           IF (#iSP <> #old.SP // SP has changed.
               OR #RTIRG_auto.Q // Auto has just been enabled, and the valve is out of pos.
               (* *)AND ABS(#iSP - #io.in.pos) > #conf.regModeMinOffset
               OR NOT #iMan AND ( // In auto
               (* *)#RTIRG_iReset.Q // Avoid dead lock
               (* *)OR #RTRIG_iFailSafe_released.Q
               (* *)OR #RTRIG_iInterlook_released.Q
               (* *)OR #RTRIG_jogClose_released.Q OR #RTRIG_jogOpen_released.Q )
               (* *)) AND (
               (*     *)NOT #iRegMode // Not regMode, no aditional requirements.
               (*     *)OR #TON_regModeWait.Q AND ( // A break between each move.
               (*        *)// Offset is bigger then a certain offset.
               (*        *)ABS(#iSP - #io.in.pos) > #conf.regModeMinOffset
               (*        *)// At almost closed and open, the offset requirement
               (*        *)// may not be fulfilled.
               (*        *)OR #io.in.pos > #conf.fullyOpenPosLim - #conf.endPosWithoutPreStop
               (*        *)OR #io.in.pos < #conf.endPosWithoutPreStop))
               // regMode should be used when a valve is controlled by a PID.
               // When the valve is in regMode, then there will be a time break between each 
               // movment. And there is a need a certain offset before an ajustment is done.
               // This behavior significantly prevents wear on the valve. If the valve is not
               // in regMode, then each change in SP will make the valve operate.
           THEN
               IF #iSP > #io.in.pos THEN
                   #action := #OPEN;
               ELSIF #iSP < #io.in.pos THEN
                   #action := #CLOSE;
               END_IF;
           END_IF;

           // --------------------------------------
           // SP-reached-pos:
           // 
           // In the main area where the valve operate, it will shut off the outputs, a
           // tiny bit before it reach the SP. This make the valve, stop exacly on SP.
           // In the area of almost closed and almost open this function is disable,
           // this makes sure that it's possible to open or close the valve entirly.
           #pre := SEL(G := #iSP > #conf.fullyOpenPosLim - #conf.endPosWithoutPreStop
                       OR #iSP < #conf.endPosWithoutPreStop,
                       IN0 := #conf.preStop, IN1 := 0);
           // Detect reached position
           IF #action = #OPEN AND (#io.in.pos > #iSP - #pre OR #io.in.fullyOpen)
               OR #action = #CLOSE AND (#io.in.pos < #iSP + #pre OR #io.in.fullyClosed)
           THEN
               #action := #NO_ACTION;
               RESET_TIMER(#TON_regModeWait);
           END_IF;
       END_IF;
       // In regMode this timer need to finnish before a new movement can be done.
       #TON_regModeWait.TON(IN := true,
                            PT := #conf.regModeTimeBreak);
   END_REGION

   REGION Gentle
       // If a big valve closes or open to fast, it can damage the pipes or other
       // equipment. This section make time breaks on closing or opening. 

       #gentleMode := #io.in.pos < #conf.gentleActivteLowLimit // ->
       // -> The function is only active under a ceratain position limit.
       AND (NOT #iFailSafe OR #conf.gentleAlsoOnFailSafe)
       // AlsoOnFailSafe: It's possible to disable the function for emergencies
       // by setting the value false.
       AND (#conf.gentleOpenEnable AND #action = #OPEN
       (* *)OR #conf.gentleCloseEnable AND #action = #CLOSE);    

       // The time break will increase as the valve move from the limit towards close.
       #pause := REAL_TO_DINT(#conf.gentleTimePauseBias
                              + (#io.in.pos / #conf.gentleActivteLowLimit)
                              * #conf.gentleTimePauseDelta);
       IF #gentleMode THEN
           #TON_gentle.TON(IN := true,
                           PT := SEL(G := #gentleAction, // Toggle times
                                     IN0 := #conf.gentleTimeRun,
                                     IN1 := #pause));
           IF #TON_gentle.Q THEN
               #gentleAction := NOT #gentleAction;
               RESET_TIMER(#TON_gentle); 
           END_IF;
           #action2 := SEL(G := #gentleAction, // Toggle action
                           IN0 := #action, IN1 := #NO_ACTION);
       ELSE
           RESET_TIMER(#TON_gentle);
           #gentleAction := false;
           // If the carefully-function is disabled, then just forward
           // the action value to the next stage.
           #action2 := #action;
       END_IF;
   END_REGION

   REGION Output
       // Make a smal time break when valve change direction. This make sure that
       // that both outputs are not active at the same time.
       #TP_toggleOut.TP(IN := #action2 <> #old.action2 AND #old.action2 <> #NO_ACTION,
                        PT := #conf.toggleTimeBreak);

       // Outputs
       IF #TP_toggleOut.Q THEN // A small time break.
           #io.out.open := false;
           #io.out.close := false;
       ELSIF #iFailSafe 
           OR #iJogClose OR #iJogOpen
       THEN
           // When failSafe or jog is active both the limit-switch and positon
           // signal most indicate that the valve is in correct position. This
           // in case one of the signals isn't working.
           #io.out.open := #action2 = #OPEN AND NOT #bothSensors.open;
           #io.out.close := #action2 = #CLOSE AND NOT #bothSensors.closed;
       ELSIF #iInterlook THEN
           #io.out.open := false;
           #io.out.close := false;
       ELSE
           #io.out.open := #action2 = #OPEN AND NOT #io.in.fullyOpen;
           #io.out.close := #action2 = #CLOSE AND NOT #io.in.fullyClosed;
       END_IF;
   END_REGION

   REGION Old    
       // Store values, to check if they has changed until next scan.
       #old.SP := #iSP;
       #old.action := #action;
       #old.action2 := #action2;
   END_REGION

   #qTimeout := #out.qucikTimeout OR #out.longTimeout;
END_FUNCTION_BLOCK

FUNCTION_BLOCK "motorValve"   // FB10, SCL
{ S7_Optimized_Access := 'TRUE' }
VERSION : 0.1
   VAR_INPUT
      iFeedbackPosition : Real;
      iFeddbackPosError : Bool;
      iFeedbackFullyOpen : Bool;
      iFeedbackFullyClosed : Bool;
   END_VAR
   VAR_OUTPUT
      qOpen : Bool;
      qClose : Bool := FALSE;
   END_VAR
   VAR RETAIN
      hmi : "motorValveHmiUdt";
   END_VAR
   VAR
      valve : "motorValveCtrl";
      SP : Real;
      SP_auto : Real;
   END_VAR
   VAR CONSTANT
      AUTO : SInt := 0;
      MAN_LOCAL : SInt := 1;
      MAN_REMOTE : SInt := 2;
   END_VAR
BEGIN
   // Valve with analog feedback.

   REGION Simulation
       IF #hmi.sim.enable AND NOT #valve.iFailSafe THEN
           // Simulation of input signal, not possible if in fail safe mode.
           #hmi.io.in.pos := #hmi.sim.pos;
           #hmi.io.in.posError := false;
           #hmi.io.in.fullyOpen := #hmi.sim.pos > #hmi.conf.fullyOpenPosLim;
           #hmi.io.in.fullyClosed := #hmi.sim.pos < #hmi.conf.fullyClosedPosLim;
       ELSE
           // Input mapping
           #hmi.io.in.pos := #iFeedbackPosition;
           #hmi.io.in.posError := #iFeddbackPosError;
           #hmi.io.in.fullyOpen := #iFeedbackFullyOpen;
           #hmi.io.in.fullyClosed := #iFeedbackFullyClosed;
       END_IF;
   END_REGION

   REGION Man / auto    
       IF #hmi.cmd.stop THEN
           #hmi.autoMan := #MAN_LOCAL;
       ELSIF #hmi.cmd.jogOpen XOR #hmi.cmd.jogClose THEN
           #hmi.autoMan := #MAN_LOCAL;
           #SP := #iFeedbackPosition;
       ELSIF #hmi.cmd.openFully XOR #hmi.cmd.closeFully THEN
           #hmi.autoMan := #MAN_LOCAL;
           #SP := SEL(G := #hmi.cmd.openFully, IN0 := 0, IN1 := 100);
       ELSIF #hmi.autoMan = #MAN_LOCAL THEN
           #SP := #hmi.SP;
       ELSIF #hmi.autoMan = #AUTO THEN
           #SP := #SP_auto;
           // If auto is controlled by a pid then #hmi.conf.regMode need to be enabled.
       END_IF;
       #hmi.SP := #valve.iSP := #SP_auto := #SP;
       // Forward auto or man to the valve controller.
       CASE #hmi.autoMan OF
           #MAN_LOCAL, #MAN_REMOTE:
               #valve.iMan := true;
           #AUTO:
               #valve.iMan := false;
       END_CASE;
   END_REGION

   REGION Valve controller.        
       // Main valve controller block.
       #valve(// iFailSafe
              // iInterlook
              // iRegMode
              iStop := #hmi.cmd.stop,
              iJogOpen := #hmi.cmd.jogOpen,
              iJogClose := #hmi.cmd.jogClose,
              iReset := #hmi.cmd.reset,
              qTimeout => #hmi.error.timeout,
              conf := #hmi.conf,
              io := #hmi.io);
       #qOpen := #hmi.io.out.open; // Outputs
       #qClose := #hmi.io.out.close;
   END_REGION

   REGION Position error    
       #hmi.error.posError :=
       #iFeedbackFullyOpen AND #iFeedbackFullyClosed
       OR #iFeedbackFullyOpen
       (* *)AND #iFeedbackPosition < #hmi.conf.fullyOpenPosLim - #hmi.conf.regModeMinOffset
       (* *)AND NOT #hmi.conf.simFullyOpenWithPos
       OR #iFeedbackFullyClosed
       (* *)AND #iFeedbackPosition > #hmi.conf.fullyClosedPosLim + #hmi.conf.regModeMinOffset
       (* *)AND NOT #hmi.conf.simFullyClosedWithPos;
   END_REGION

   REGION End
       // Count secounds the valve has been operating, and number of starts.
       "operatingTime"(in := #qOpen OR #qClose,
                       opr := #hmi.operatingTime);

       // Reset signals.
       #hmi.cmd.jogOpen := false;
       #hmi.cmd.jogClose := false;
       #hmi.cmd.openFully := false;
       #hmi.cmd.closeFully := false;
       #hmi.cmd.reset := false;
       #hmi.cmd.man := false;
       #hmi.cmd.auto := false;
       CASE #hmi.autoMan OF // Reset stop signal, only if in man.
           #MAN_LOCAL, #MAN_REMOTE: // If in auto, then do nothing.
               #hmi.cmd.stop := false;
       END_CASE;

       // Other signals to HMI
       #hmi.info.failSafe := #valve.iFailSafe;
       #hmi.info.interlook := #valve.iInterlook;
       #hmi.info.regMode := #valve.iRegMode;

       #hmi.sim.simByPlc := #hmi.io.simulated;
       #hmi.io.simulated := false;
   END_REGION
END_FUNCTION_BLOCK

FUNCTION_BLOCK "motorValveSimulation"   // FB20, SCL
{ S7_Optimized_Access := 'TRUE' }
VERSION : 0.1
   VAR_INPUT
      speed : Real := 1.0;
   END_VAR
   VAR_IN_OUT
      io : "motorValveIoUdt";
   END_VAR
   VAR
      old : UDInt;
      sn : UDInt;
   END_VAR
   VAR_TEMP
      t : DTL;
      "e" : Int;
   END_VAR
BEGIN
   #"e" := RD_SYS_T(#t);
   #sn := #t.NANOSECOND / 100000 + #t.SECOND * 10;

   IF #sn = #old THEN
       IF #io.out.open THEN
           #io.in.pos += #speed * 0.1;
       ELSIF #io.out.close THEN
           #io.in.pos -= #speed;
       END_IF;
   END_IF;
   #old := #sn;

   #io.in.pos := LIMIT(MN := 0, IN := #io.in.pos, MX := 100);
   #io.in.fullyOpen := #io.in.pos > 99;
   #io.in.fullyClosed := #io.in.pos < 1;

   #io.simulated := true;
END_FUNCTION_BLOCK

// folder: _ state macine

FUNCTION_BLOCK "stateMachineTimer"   // FB1, SCL
{ S7_Optimized_Access := 'TRUE' }
VERSION : 0.1
   VAR_INPUT
      state : Int;   // state machine
   END_VAR
   VAR_OUTPUT
      q : Bool;   // out
      rt : Time;   // Remaining time
      et : Time;
   END_VAR
   VAR
      pt : Time;   // input time
      "timer" : IEC_TIMER;
      old_state : Int;
   END_VAR
BEGIN
   // https://github.com/rexhip/
   //
   // State machine timer.
   // 
   // The timer is reseted if:
   // - Pt hasen't got a new value (for each scan)
   // - New state

   #"timer".TON(IN := #pt <> T#0s
              (* *)AND #state = #old_state,
              PT := #pt,
              Q => #q);

   #et := #"timer".ET;
   #rt := #pt - #et;

   #pt := T#0s;
   #old_state := #state;
END_FUNCTION_BLOCK

FUNCTION_BLOCK "setResetTimer"   // FB3, SCL
{ S7_Optimized_Access := 'TRUE' }
VERSION : 0.1
   VAR_INPUT
      in : Bool;
      pt : Time;
      set : Bool;
      reset : Bool;
   END_VAR
   VAR_OUTPUT
      q : Bool;
   END_VAR
   VAR
      "timer" : IEC_TIMER;
      timer_q : Bool;
   END_VAR
BEGIN
   // Once the timer has elapsed, the output
   // will stay true until it's reset.

   #"timer".TON(IN := #in, PT := #pt, Q => #timer_q);

   IF #set THEN
       #q := true;
   ELSIF #reset THEN
       #q := false;
   ELSIF #timer_q THEN
       #q := true;
   END_IF;
END_FUNCTION_BLOCK

FUNCTION "sTimer" : Bool   // FC2, SCL
{ S7_Optimized_Access := 'TRUE' }
VERSION : 0.1
   VAR_INPUT
      pt : Time;
   END_VAR
   VAR_IN_OUT
      t : "stateMachineTimer";
   END_VAR
BEGIN
   // sTimer
   // Make a timer, a one liner, in a state macine

   #t.pt := #pt;
   #sTimer := #t.q;
END_FUNCTION

// folder: io

FUNCTION_BLOCK "ioGlobal_FB"   // FB1, SCL
{ S7_Optimized_Access := 'TRUE' }
VERSION : 0.1
   VAR
      hmi : "ioGlobalUdt";
      z_internal_timer : IEC_TIMER;
      z_internal : Struct
         fs : Bool := TRUE;
         timer_mem : Time;
      END_STRUCT;
      collectInfo : Struct
         activeSimCnt : UInt;
         activeAlarmsCnt : UInt;
         unacknowledgedAlarmsCnt : UInt;
         errorCnt : UInt;
      END_STRUCT;
      info2ioBlocks : Struct
         runtimeDiff : Time;
         ackAllAlarms : Bool;
         disableAllSim : Bool;
         firstScan : Bool := TRUE;
      END_STRUCT;
      z : Struct
         ioIdCnt : UInt;
      END_STRUCT;
      copyPaste : "analogInAndAlarmsUdt";
      normX : "normXAnalogUdt";
   END_VAR
BEGIN
   // ioGlobal: This block handels common function for io, eg:
   //  - Count active simulations
   //  - Disable all simulations
   //  - Count active alarms
   //  - Ack. all active alarms

   // Calculate time of each plc scan.
   #z_internal_timer.TON(IN := NOT #z_internal_timer.Q, PT := T#24d);
   IF #z_internal_timer.ET <> #z_internal.timer_mem THEN
       #info2ioBlocks.runtimeDiff := #z_internal_timer.ET - #z_internal.timer_mem;
   END_IF;
   #z_internal.timer_mem := #z_internal_timer.ET;

   // First scan
   #info2ioBlocks.firstScan := #z_internal.fs;
   #z_internal.fs := false;

   // Common information to all io-blocks.
   #info2ioBlocks.ackAllAlarms := #hmi.ackAllAlarms;
   #info2ioBlocks.disableAllSim := #hmi.disableAllSim;
   // Make sure that ack only happens once.
   #hmi.ackAllAlarms := false;
   #hmi.disableAllSim := false;

   // Information from io-blocks.
   #hmi.totalActiveAlarms := #collectInfo.activeAlarmsCnt;
   #hmi.totalActiveSim := #collectInfo.activeSimCnt;
   #hmi.totalUnacknowledgedAlarms := #collectInfo.unacknowledgedAlarmsCnt;
   #hmi.totalErrors := #collectInfo.errorCnt;
   // Reset the counter for new collection of info on next scan.
   #collectInfo.activeAlarmsCnt := 0;
   #collectInfo.activeSimCnt := 0;
   #collectInfo.unacknowledgedAlarmsCnt := 0;
   #collectInfo.errorCnt := 0;

   // ioId io-id
   #z.ioIdCnt := 0;

   // ( https://github.com/rexhip/ )
END_FUNCTION_BLOCK

FUNCTION "alarmReal" : Void   // FC2, SCL
{ S7_Optimized_Access := 'TRUE' }
VERSION : 0.1
   VAR_INPUT
      value : Real;   // Value that will be compared
      action : SInt;   // 1=Greater then, 2=less then
      disable : Bool;   // diable alarm
   END_VAR
   VAR_IN_OUT
      runtimeDiff : Time;   // Time of last program scan, used for internal timer
      alarm : "alarmRealUdt";
   END_VAR
   VAR_TEMP
      tmpQset : Bool;
      tmpQrst : Bool;
   END_VAR
   VAR CONSTANT
      LESS_THEN : SInt := 1;
      GREATER_THEN : SInt := 2;
   END_VAR
BEGIN
   // Value alarm

   #alarm.value := #value;
   #alarm.action := #action;

   IF #alarm.enable AND NOT #disable THEN
       CASE #action OF
           #LESS_THEN: // (1)
               #tmpQset := #value < #alarm.lim;
               #tmpQrst := #value > #alarm.lim + #alarm.hyst;
           #GREATER_THEN: // (2)
               #tmpQset := #value > #alarm.lim;
               #tmpQrst := #value < #alarm.lim - #alarm.hyst;
       END_CASE;
       IF #alarm.Q THEN  // if alarm has been activated.
           #alarm.memAck := #alarm.memAck OR #alarm.ack; // Acknowledge
           IF #tmpQrst AND (
               #alarm.autoAck
               OR #alarm.memAck AND NOT #alarm.dobleAck
               OR #alarm.ack AND #alarm.dobleAck)
           THEN
               #alarm.Q := false;
           END_IF;
       ELSE  // Not #alarm.Q
           IF #tmpQset THEN
               #alarm.delayEt += #runtimeDiff;
               IF #alarm.delayEt >= #alarm.delay THEN
                   #alarm.Q := true;
                   #alarm.memAck := false;
               END_IF;
           ELSE
               #alarm.delayEt := T#0s;
           END_IF;
       END_IF;
       #alarm.ack := false;

   ELSE // Alarm disabled
       #alarm.Q := false;
       #alarm.delayEt := T#0s;
   END_IF;

   // ( https://github.com/rexhip/ )
END_FUNCTION

FUNCTION "ioGlobalAlarmLinking" : Void   // FC3, SCL
{ S7_Optimized_Access := 'TRUE' }
VERSION : 0.1
   VAR_IN_OUT
      alarm : "alarmRealUdt";
      ioGlobal : "ioGlobal_FB";
   END_VAR
BEGIN
   // Connecting ioGlobal functions with valueAlarm.

   // Acknowle alarm
   #alarm.ack := #ioGlobal.info2ioBlocks.ackAllAlarms;

   // Count active alarms
   #ioGlobal.collectInfo.activeAlarmsCnt += BOOL_TO_UINT(#alarm.Q);
   // Count unacknowledged alarms
   #ioGlobal.collectInfo.unacknowledgedAlarmsCnt +=
   BOOL_TO_UINT(#alarm.Q AND NOT #alarm.memAck);

   // ( https://github.com/rexhip/ )
END_FUNCTION

FUNCTION "alarmBoolSimple" : Void   // FC5, SCL
{ S7_Optimized_Access := 'TRUE' }
VERSION : 0.1
   VAR_INPUT
      in : Bool;
   END_VAR
   VAR_IN_OUT
      alarm : "alarmBoolSimpleUdt";
   END_VAR
BEGIN
   // Simple digital alarm 

   IF #alarm.enable THEN
       IF #alarm.Q THEN
           #alarm.memAck := #alarm.memAck OR #alarm.ack; // Acknowledge
           IF NOT #alarm.in AND (
               #alarm.autoAck
               OR #alarm.memAck AND NOT #alarm.dobleAck
               OR #alarm.ack AND #alarm.dobleAck)
           THEN
               #alarm.Q := false;
           END_IF;
       ELSIF #alarm.in THEN
           #alarm.Q := true;
           #alarm.memAck := false;
       END_IF;
       #alarm.ack := false;

   ELSE // Alarm is disabled
       #alarm.Q := false;
   END_IF;
END_FUNCTION

FUNCTION "digitalOut" : Void   // FC8, SCL
{ S7_Optimized_Access := 'TRUE' }
VERSION : 0.1
   VAR_OUTPUT
      Out : Bool;
   END_VAR
   VAR_IN_OUT
      doUdt : "digitalOutUdt";
      ioGlobal : "ioGlobal_FB";
   END_VAR
   VAR_TEMP
      t : Bool;
   END_VAR
BEGIN
   // Digital out
   //
   // - For most application a analog output block is not needed. However
   //
   // - failSafe: Output will go to a predefined value set by failSafeValue (%),
   //   this can be used for emergency stop, simulation will not work when
   //   failSafe is activated.

   // A id for each io
   #ioGlobal.z.ioIdCnt += 1;

   IF #doUdt.disableSim OR #ioGlobal.info2ioBlocks.disableAllSim THEN
       #doUdt.simEnable := false;
   END_IF;

   IF #doUdt.failSafe THEN
       #t := #doUdt.failSafeValue;
   ELSE
       #t := SEL(G := #doUdt.simEnable,
                 IN0 := #doUdt.in XOR #doUdt.invert,
                 IN1 := #doUdt.simValue);
   END_IF;
   #doUdt.simValue := #Out := #t;

   #ioGlobal.collectInfo.activeSimCnt += BOOL_TO_USINT(#doUdt.simEnable);

   // ( https://github.com/rexhip/ )
END_FUNCTION

FUNCTION "digitalIn" : Void   // FC10, SCL
{ S7_Optimized_Access := 'TRUE' }
VERSION : 0.1
   VAR_INPUT
      in : Bool;
   END_VAR
   VAR_IN_OUT
      diUdt : "digitalInUdt";
      ioGlobal : "ioGlobal_FB";
   END_VAR
   VAR_TEMP
      "e" : Int;
      tmpQ : Bool;
      tmpIn : Bool;
   END_VAR
BEGIN
   // Digital input ( https://github.com/rexhip/ )

   // A id for each io
   #ioGlobal.z.ioIdCnt += 1;

   IF #diUdt.sim THEN
       #diUdt.delayEt := T#0ms;
   ELSE
       #tmpQ := #diUdt.Q;
       #tmpIn := #in XOR #diUdt.invert;
       IF #tmpIn AND NOT #diUdt.Q THEN
           #diUdt.delayEt += #ioGlobal.info2ioBlocks.runtimeDiff;
       ELSIF NOT #tmpIn THEN
           #diUdt.delayEt := T#0ms;
       END_IF;
       #diUdt.Q := #diUdt.delayEt >= #diUdt.delay;

       // Logging - the time the input change state.
       IF #diUdt.Q AND NOT #tmpQ THEN
           #"e" := RD_LOC_T(#diUdt.timeOn);
       ELSIF NOT #diUdt.Q AND #tmpQ THEN
           #"e" := RD_LOC_T(#diUdt.timeOff);
       END_IF;
   END_IF;

   "alarmBoolSimple"(in := #diUdt.Q, alarm := #diUdt.alarm);

   // Count alarms, errors and simulations.
   #ioGlobal.collectInfo.activeAlarmsCnt += BOOL_TO_UINT(#diUdt.alarm.Q);
   #ioGlobal.collectInfo.errorCnt += BOOL_TO_UINT(#diUdt.Error);;
   #ioGlobal.collectInfo.activeSimCnt += BOOL_TO_UINT(#diUdt.sim);

   // ( https://github.com/rexhip/ )
END_FUNCTION

FUNCTION "analogInError" : Bool   // FC14, SCL
{ S7_Optimized_Access := 'TRUE' }
VERSION : 0.1
   VAR_INPUT
      in : Int;
   END_VAR
   VAR_TEMP
      t : Real;
   END_VAR
BEGIN
   // Analog in error (outside limits.)
   #analogInError := #in < -4864 OR #in > 32512;;
END_FUNCTION

FUNCTION "syncReal" : Void   // FC17, SCL
{ S7_Optimized_Access := 'TRUE' }
VERSION : 0.1
   VAR_IN_OUT
      prim : Real;   // primary
      sec : Real;   // secoundary
      memory : Real;
   END_VAR
BEGIN
   // Make two variables have the same value. If one change, the
   // value will be transfer to the other one.

   IF #prim = #memory THEN
       #prim := #sec;
   ELSE
       #sec := #prim;
   END_IF;

   #memory := #sec;
END_FUNCTION

FUNCTION "setUnipolar" : Void   // FC18, SCL
{ S7_Optimized_Access := 'TRUE' }
VERSION : 0.1
   VAR_IN_OUT
      unipolar : "normXAnalogUdt";
   END_VAR
BEGIN
   // Set values for analog input and output to
   // unipolar.

   #unipolar.rawMin := 0;
   #unipolar.rawMax := 27648;

   // Outside limits bellow will generate error.
   #unipolar.errorLimMin := -4864;
   #unipolar.errorLimMax := 32512;
END_FUNCTION

FUNCTION "setAnalogType" : "normXAnalogUdt"   // FC19, SCL
{ S7_Optimized_Access := 'TRUE' }
VERSION : 0.1
   VAR_INPUT
      select : Int;
   END_VAR
   VAR_TEMP
      dommy : "normXAnalogUdt";
   END_VAR
BEGIN
   // Set values for analog input and output 

   CASE #select OF
       1:  // Siemens unipolar
           #setAnalogType.rawMin := 0;
           #setAnalogType.rawMax := 27648;
           #setAnalogType.errorLimMin := -4864;
           #setAnalogType.errorLimMax := 32512;
       2:  // Siemens bipolar
           #setAnalogType.rawMin := -27648;
           #setAnalogType.rawMax := 27648;
           #setAnalogType.errorLimMin := -32512;
           #setAnalogType.errorLimMax := 32512;
       3:  // Wago - 750-496  - 0/4-20 mA
           #setAnalogType.rawMin := 0;
           #setAnalogType.rawMax := 30832;
           #setAnalogType.errorLimMin := -773;
           #setAnalogType.errorLimMax := 32763;
           // 4:  
           //  #setAnalogType.min := ;
           //  #setAnalogType.max := ;
           //  #setAnalogType.errorLimMin := ;
           //  #setAnalogType.errorLimMax := ;
       ELSE
           #setAnalogType := #dommy;
   END_CASE;
END_FUNCTION

FUNCTION "pasteAnalogInSetting" : Void   // FC20, SCL
{ S7_Optimized_Access := 'TRUE' }
VERSION : 0.1
   VAR_IN_OUT
      src : "analogInAndAlarmsUdt";
      dest : "analogInAndAlarmsUdt";
   END_VAR
BEGIN
   // Select only the settings and not values from the 
   // udt's and transfer them from src to dest.

   #dest.ai.offset := #src.ai.offset ;
   #dest.ai.errorAction := #src.ai.errorAction ;
   #dest.ai.gain := #src.ai.gain ;
   #dest.ai.filterConst := #src.ai.filterConst ;
   #dest.ai.forceInsideScale := #src.ai.forceInsideScale ;
   #dest.ai.scaleMax := #src.ai.scaleMax ;
   #dest.ai.scaleMin := #src.ai.scaleMin ;

   "pasteAlarmSetting"(src := #src.alarmHH, dest := #dest.alarmHH);
   "pasteAlarmSetting"(src := #src.alarmH,  dest := #dest.alarmH);
   "pasteAlarmSetting"(src := #src.alarmLL, dest := #dest.alarmLL);
   "pasteAlarmSetting"(src := #src.alarmL,  dest := #dest.alarmL);
END_FUNCTION

FUNCTION "pasteAlarmSetting" : Void   // FC21, SCL
{ S7_Optimized_Access := 'TRUE' }
VERSION : 0.1
   VAR_IN_OUT
      src : "alarmRealUdt";
      dest : "alarmRealUdt";
   END_VAR
BEGIN

   #dest.enable := #src.enable;
   #dest.autoAck := #src.autoAck ;
   #dest.delay := #src.delay ;
   #dest.hyst := #src.hyst ;
   #dest.lim := #src.lim ;
END_FUNCTION

FUNCTION "analogOutSimple" : Int   // FC22, SCL
{ S7_Optimized_Access := 'TRUE' }
VERSION : 0.1
   VAR_INPUT
      in : Real;   // Percent
   END_VAR
   VAR_TEMP
      x : Real;
   END_VAR
BEGIN
   // Simple analog unipolar output

   // Input:  per cent.
   // Output: Siemens unipolar scale.

   #x := LIMIT(MN := 0, IN := #in / 100, MX := 1);
   #analogOutSimple := SCALE_X(MIN := 0, VALUE := #x, MAX := 27648);

   // ( https://github.com/rexhip/ )
END_FUNCTION

FUNCTION "syncBool" : Void   // FC27, SCL
{ S7_Optimized_Access := 'TRUE' }
VERSION : 0.1
   VAR_IN_OUT
      prim : Bool;   // primary
      sec : Bool;   // secoundary
      memory : Bool;
   END_VAR
BEGIN
   // Make two variables have the same value. If one change, the
   // value will be transfer to the other one.

   IF #prim = #memory THEN
       #prim := #sec;
   ELSE
       #sec := #prim;
   END_IF;

   #memory := #sec;
END_FUNCTION

// folder: io/example

FUNCTION_BLOCK "_example_analogOutpus"   // FB2, SCL
{ S7_Optimized_Access := 'TRUE' }
VERSION : 0.1
   VAR_OUTPUT
      ao_FV01 : Int;
      ao_FV02 : Int;
      ao_FV03 : Int;
   END_VAR
   VAR_IN_OUT
      ioGlobal : "ioGlobal_FB";
   END_VAR
   VAR RETAIN
      FV01 : "analogOutUdt";
      FV02 : "analogOutUdt";
   END_VAR
   VAR
      FV03 : Real;
   END_VAR
BEGIN


   "analogOut"(aoUdt := #FV01,
               ioGlobal := #ioGlobal,
               q => #ao_FV01);

   "analogOut"(aoUdt := #FV02,
               ioGlobal := #ioGlobal,
               q => #ao_FV02);

   // Very simple analog output.
   #ao_FV03 := "analogOutSimple"(#FV03);
END_FUNCTION_BLOCK

FUNCTION_BLOCK "_example_digitalInputs"   // FB3, SCL
{ S7_Optimized_Access := 'TRUE' }
VERSION : 0.1
   VAR_INPUT
      di_PAH01 : Bool;
      di_PAH02 : Bool;
   END_VAR
   VAR_IN_OUT
      ioGlobal : "ioGlobal_FB";
   END_VAR
   VAR RETAIN
      PAH01 : "digitalInUdt";
      PAH02 : "digitalInUdt";
   END_VAR
BEGIN

   "digitalIn"(in := #di_PAH01,
               diUdt := #PAH01,
               ioGlobal := #ioGlobal);
   "digitalIn"(in := #di_PAH02,
               diUdt := #PAH02,
               ioGlobal := #ioGlobal);
END_FUNCTION_BLOCK

FUNCTION_BLOCK "_example_digitalOutpus"   // FB4, SCL
{ S7_Optimized_Access := 'TRUE' }
VERSION : 0.1
   VAR_OUTPUT
      do_PX01 : Bool;
      do_PX02 : Bool;
   END_VAR
   VAR_IN_OUT
      ioGlobal : "ioGlobal_FB";
   END_VAR
   VAR RETAIN
      PX01 : "digitalOutUdt";
      PX02 : "digitalOutUdt";
   END_VAR
BEGIN

   "digitalOut"(Out => #do_PX01,
                doUdt := #PX01,
                ioGlobal := #ioGlobal);

   "digitalOut"(Out => #do_PX02,
                doUdt := #PX02,
                ioGlobal := #ioGlobal);
END_FUNCTION_BLOCK

FUNCTION_BLOCK "_example_analogInputs"   // FB5, SCL
{ S7_Optimized_Access := 'TRUE' }
VERSION : 0.1
   VAR_INPUT
      ai_FT12 : Int;
      ai_TT27 : Int;
      value_from_other_source : Real;
   END_VAR
   VAR_IN_OUT
      ioGlobal : "ioGlobal_FB";
   END_VAR
   VAR RETAIN
      FT12 : "analogInAndAlarmsUdt";
      TT27 : "analogInAndAlarmsUdt";
      PT44 : "analogInAndAlarmsUdt";
   END_VAR
BEGIN
   // Analog inputs example. ( https://github.com/rexhip/ )

   // In a real world example the input on this block
   // would be PLC-tags connected to fysical IO.

   "analogInAndAlarms"(in := #ai_FT12,
                       aiUdt := #FT12,
                       ioGlobal := #ioGlobal);
   "analogInAndAlarms"(in := #ai_TT27,
                       aiUdt := #TT27,
                       ioGlobal := #ioGlobal);

   // Value arriving from other source, eg. profinet.
   "analogInReal"(in := #value_from_other_source,
                  error := false, // Should be provided in case comm. error.
                  aiUdt := #PT44,
                  ioGlobal := #ioGlobal);
END_FUNCTION_BLOCK

// folder: io/hmi multiplex

FUNCTION "syncAlarmReal" : Void   // FC26, SCL
{ S7_Optimized_Access := 'TRUE' }
VERSION : 0.1
   VAR_IN_OUT
      prim : "alarmRealUdt";
      sec : "alarmRealUdt";
      memory : "alarmRealUdt";
   END_VAR
BEGIN

   #prim.value := #sec.value;
   #prim.action := #sec.action;

   "syncReal"(prim := #prim.lim ,
              sec := #sec.lim ,
              memory := #memory.lim);

   "syncBool"(prim := #prim.Q,
              sec := #sec.Q,
              memory := #memory.Q);
END_FUNCTION

// folder: motor valve

FUNCTION "operatingTime" : Void   // FC12, SCL
{ S7_Optimized_Access := 'TRUE' }
VERSION : 0.1
   VAR_INPUT
      in : Bool;
   END_VAR
   VAR_IN_OUT
      opr : "operatingTimeUdt";
   END_VAR
   VAR_TEMP
      "e" : Int;
      rdSysT : DTL;
   END_VAR
BEGIN
   // This function shouldn't be used with periodical interupts that has longer
   // cycles then 50 secounds.

   // Operating time.
   // (Max value: 2^32 / (24 * 60*60 * 365) = 136 => 136 years.)
   #"e" := RD_SYS_T(#rdSysT);
   #opr.operatingTime +=
   SEL(G := #in, IN0 := 0, IN1 := (#rdSysT.SECOND - #opr.oldSec + 60) MOD 60);
   #opr.oldSec := #rdSysT.SECOND;

   // Start cnt.
   #opr.startCnt += BOOL_TO_UDINT(#in AND NOT #opr.oldIn);
   #opr.oldIn := #in;
END_FUNCTION

FUNCTION "time_to_real" : Real   // FC28, SCL
{ S7_Optimized_Access := 'TRUE' }
VERSION : 0.1
   VAR_INPUT
      in : Time;
   END_VAR
BEGIN

   #time_to_real := DINT_TO_REAL(T_CONV( #in)) / 1000;
END_FUNCTION

// folder: pid

FUNCTION_BLOCK "pid"   // FB19, SCL
{ S7_Optimized_Access := 'TRUE' }
VERSION : 0.1
   VAR
      pidUdt : "pidUdt";
      pidCompact : PID_Compact;
      oldSec : USInt;
   END_VAR
   VAR_TEMP
      T : DTL;
      "e" : Int;
   END_VAR
BEGIN


   #"e" := RD_SYS_T(#T);
   IF #T.SECOND <> #oldSec THEN
       #pidCompact.Retain.CtrlParams := #pidUdt.pidParam;
       #pidCompact(Setpoint := #pidUdt.sp,
                   Input := #pidUdt.pv,
                   ManualEnable := #pidUdt.man,
                   Output => #pidUdt.mv,
                   Error => #pidUdt.error);
   END_IF;
   #oldSec := #T.SECOND;
END_FUNCTION_BLOCK

// folder: sr

FUNCTION "setReset_rd" : Void   // FC15, SCL
{ S7_Optimized_Access := 'TRUE' }
VERSION : 0.1
   VAR_INPUT
      s : Bool;
      r : Bool;
   END_VAR
   VAR_IN_OUT
      q : Bool;
   END_VAR
BEGIN
   // Set-reset (sd = reset dominant)

   IF #r THEN
       #q := false;
   ELSIF #s THEN
       #q := true;
   END_IF;
END_FUNCTION

FUNCTION "setReset_sd" : Void   // FC16, SCL
{ S7_Optimized_Access := 'TRUE' }
VERSION : 0.1
   VAR_INPUT
      s : Bool;
      r : Bool;
   END_VAR
   VAR_IN_OUT
      q : Bool;
   END_VAR
BEGIN
   // Set-reset (sd = reset dominant)

   IF #s THEN
       #q := true;
   ELSIF #r THEN
       #q := false;
   END_IF;
END_FUNCTION

// folder: zSlib/misc/conv/time_to_str

FUNCTION "str::" : String   // FC29, SCL
{ S7_Optimized_Access := 'TRUE' }
VERSION : 0.1
   VAR_INPUT
      in : Time;   // Time to be converted in to string.
   END_VAR
   VAR_TEMP
      t : DTL;
      dayOrHour : Bool;
   END_VAR
BEGIN
   // Time to string.

   #t += #in; // Implicit convert to dtl.
   #t.DAY -= 1; 
   #time_to_str := ''; // (Avoiding compilation warnings) 

   IF #t.DAY <> 0 THEN
       #time_to_str := CONCAT(IN1 := RIGHT
                              (IN := S_CONV(#t.DAY),
                               L := 1 + BOOL_TO_INT(#t.DAY > 9)),
                              IN2 := ', ');
   END_IF;
   IF #t.HOUR <> 0 OR LEN(#time_to_str) <> 0 THEN
       #time_to_str := CONCAT(IN1 := #time_to_str,
                              IN2 := RIGHT
                              (IN := S_CONV(#t.HOUR),
                               L := 1 + BOOL_TO_INT(#t.HOUR > 9)),
                              IN3 := ':');
   END_IF;
   #time_to_str := CONCAT(IN1 := #time_to_str,
                          IN2 := RIGHT
                          (IN := S_CONV(#t.MINUTE),
                           L := 1 + BOOL_TO_INT(#t.MINUTE > 9)),
                          IN3 := ':');
   #time_to_str := CONCAT(IN1 := #time_to_str,
                          IN2 := RIGHT
                          (IN := S_CONV(#t.SECOND),
                           L := 1 + BOOL_TO_INT(#t.SECOND > 9)));

   // https://github.com/rexhip/
END_FUNCTION

// ===== library: MasterCopy "ponselMessure_ChangeMbAddr" =====

FUNCTION_BLOCK "ponselMessure_ChangeMbAddr"   // FB2, SCL
{ S7_Optimized_Access := 'TRUE' }
VERSION : 0.1
   VAR_INPUT
      current_addr : USInt;
      new_addr : UInt;
      exec : Bool := true;
   END_VAR
   VAR_OUTPUT
      Done : Bool;
      Error : Bool;
   END_VAR
   VAR_IN_OUT
      mb_query : "mb_query";
   END_VAR
   VAR_TEMP
      d : Bool;
      "e" : Bool;
   END_VAR
BEGIN
   IF #new_addr < 1 OR #new_addr > 247
       OR #new_addr = #current_addr
   THEN
       #"e" := TRUE;
   ELSIF #exec THEN
       #mb_query(mb_addr := #current_addr,
                 mode := #mb_query.c.write.holding_reg,
                 data_addr := 16#A3,
                 Done => #d,
                 Error => #"e",
                 data_ptr := #new_addr);
   END_IF;
   #Done := #d;
   #Error := #"e";
END_FUNCTION_BLOCK

// ===== library: MasterCopy "ponselMessure_changeParity" =====

FUNCTION_BLOCK "ponselMessure_changeParity"   // FB9, SCL
{ S7_Optimized_Access := 'TRUE' }
VERSION : 0.1
   VAR_INPUT
      mb_addr : USInt;
      parity : USInt;
   END_VAR
   VAR_OUTPUT
      Done : Bool;
      Error : Bool;
   END_VAR
   VAR_IN_OUT
      mb_query : "mb_query";
   END_VAR
   VAR_TEMP
      d : Bool;
      "e" : Bool;
      "word" : Word;
   END_VAR
BEGIN
   // This block isn't finnish.
   //
   IF #parity > 3 THEN
       #"e" := TRUE;
   ELSE
       CASE #parity OF
           0:  // None
               #"word".%X0 := false;
               #"word".%X1 := false;
           1:  // Odd
               #"word".%X0 := false;
               #"word".%X1 := true;
           2:  // Even
               #"word".%X0 := true;
               #"word".%X1 := false;
       END_CASE;
       (*#mb_query(mb_addr := #mb_addr,
                 mode := #mb_query.c.write.holding_reg,
                 data_addr := ,
                 Done => #d,
                 Error => #e,
                 data_ptr := #word);*)
   END_IF;
   #Done := #d;
   #Error := #"e";
END_FUNCTION_BLOCK

// ===== library: MasterCopy "ponselMessure_readSign" =====

FUNCTION_BLOCK "ponselMessure_readSign"   // FB8, SCL
{ S7_Optimized_Access := 'TRUE' }
VERSION : 0.1
   VAR_INPUT
      mb_addr : USInt;
   END_VAR
   VAR_OUTPUT
      Done : Bool;
      Error : Bool;
   END_VAR
   VAR_IN_OUT
      mb_query : "mb_query";
   END_VAR
   VAR
      signs : Array[1..3] of String[64];
   END_VAR
BEGIN
   // Read calibration signatures

   #mb_query(mb_addr := #mb_addr,
             mode := #mb_query.c.read.holding_reg,
             data_addr := 16#027e,
             data_ptr := #signs);

   IF #mb_query.Done THEN
       #Done := true;
       #Error := false;
   ELSIF #mb_query.Error THEN
       #Done := false;
       #Error := true;
   END_IF;
END_FUNCTION_BLOCK

// ===== library: MasterCopy "ponselMessure_readUnits" =====

FUNCTION_BLOCK "ponselMessure_readUnits"   // FB2, SCL
{ S7_Optimized_Access := 'TRUE' }
VERSION : 0.1
   VAR_INPUT
      mb_addr : USInt;
   END_VAR
   VAR_OUTPUT
      Done : Bool;
      Error : Bool;
   END_VAR
   VAR_IN_OUT
      mb_query : "mb_query";
   END_VAR
   VAR
      Units : Array[0..4] of String[6];
   END_VAR
BEGIN
   // 

   #mb_query(mb_addr := #mb_addr,
             mode := #mb_query.c.read.holding_reg,
             data_addr := 16#0D22,
             data_ptr := #Units);
   IF #mb_query.Done THEN
       #Done := true;
       #Error := false;
   ELSIF #mb_query.Error THEN
       #Done := false;
       #Error := true;
   END_IF;
END_FUNCTION_BLOCK

// ===== library: MasterCopy "ponselMessure_restoreDefaultCoefficients" =====

FUNCTION_BLOCK "ponselMessure_restoreDefaultCoefficients"   // FB2, SCL
{ S7_Optimized_Access := 'TRUE' }
VERSION : 0.1
   VAR_INPUT
      mb_addr : USInt;
      restorTemp : Bool;
      restorPar1 : Bool;
      restorPar2 : Bool;
      restorPar3 : Bool;
      restorPar4 : Bool;
   END_VAR
   VAR_OUTPUT
      Done : Bool;
      Error : Bool;
   END_VAR
   VAR_IN_OUT
      mb_query : "mb_query";
   END_VAR
   VAR
      "word" : Word;
      old_word : Word;
      first_scan : Bool := true;
   END_VAR
   VAR_TEMP
      d : Bool;
      "e" : Bool;
   END_VAR
BEGIN
   // Restore default calibration coefficients.

   #"word".%X0 := #restorTemp;
   #"word".%X1 := #restorPar1;
   #"word".%X2 := #restorPar2;
   #"word".%X3 := #restorPar3;
   #"word".%X4 := #restorPar4;

   IF #"word" <> #old_word AND NOT #first_scan THEN
       #mb_query(mb_addr := #mb_addr,
                 mode := #mb_query.c.write.holding_reg,
                 data_addr := 16#02,
                 Done => #d,
                 Error => #"e",
                 data_ptr := #"word");
   END_IF;
   #old_word := #"word";

   #first_scan := false;
   #Done := #d;
   #Error := #"e";
END_FUNCTION_BLOCK

// ===== library: MasterCopy "ponselMesure_calibrate" =====

FUNCTION_BLOCK "ponselMesure_calibrate"   // FB5, SCL
{ S7_Optimized_Access := 'TRUE' }
VERSION : 0.1
   VAR_INPUT
      ref_value : Real;
   END_VAR
   VAR_OUTPUT
      Done : Bool;
      Error : Bool;
   END_VAR
   VAR_IN_OUT
      mb_query : "mb_query";
      ponsel_messure : "Ponsel_mesure";
      sign : "ponselMesure_sign_udt";
   END_VAR
   VAR
      conf : Struct
         messurementsBeforeCal : USInt;
      END_STRUCT;
      mode : USInt;
      state : Int;
      oldQueryCnt : UDInt;
      error_cnt : USInt;
      dword_14c : DWord;
   END_VAR
   VAR_TEMP
      valid_value : Bool;
      tDword : DWord;
      empty : "ponselMesure_sign_udt";
   END_VAR
BEGIN
   #mb_query.mb_addr := #ponsel_messure.mb_addr;
   #mb_query.mode := #mb_query.c.write.holding_reg;
   #mb_query.Error := false;

   #Done := false;
   #Error := false;

   CASE #state OF

       10: // Wait for start signal
           #state += 1;
           #oldQueryCnt := #ponsel_messure.QueryCnt;

       11: // Do some messurements.
           #ponsel_messure.api.interval := T#2s;
           #state += BOOL_TO_INT(#ponsel_messure.QueryCnt - #oldQueryCnt >
                                 #conf.messurementsBeforeCal
                                 AND #ponsel_messure.Measurement_ok);
           #state := SEL(G := #mode = 0, IN0 := #state, IN1 := 0);
       12: // Stop messurement
           #ponsel_messure.api.wait := true;
           #state += BOOL_TO_INT(#ponsel_messure.api.idle);
       13: // Send ref. value to transmitter
           #ponsel_messure.api.wait := true; // stop messurement.
           CASE #mode OF
               1..10: // Parameters, 1 to 10
                   #mb_query.data_addr := 16#204 + (#mode - 1) * 2;
               11..12: // Temperature.
                   #mb_query.data_addr := 16#200 + (#mode - 11) * 2;
           END_CASE;
           #mb_query(data_ptr := #ref_value);
           #state += BOOL_TO_INT(#mb_query.Done);
       14: // Preperation for 14c, the word may be later written to device.
           CASE #mode OF
               1..4: // Parameter, 1 - 4  
                   #tDword.%X2 := true;
                   #tDword := SHL(IN := #tDword, N := #mode - 1);
               11: // Temperature zero and span.
                   #tDword.%X0 := true;
                   #tDword := SHL(IN := #tDword, N := #mode - 11);
           END_CASE;
           #dword_14c := #dword_14c OR #tDword; // A the bit "14c"
           #state += 1;

           // =============
           // Save

       20: // Send signature to transmitter.
           CASE #mode OF
               1..4: // Parameter, 1 - 4  // ( 16#28e - 16#27e = 16#10 )
                   #mb_query.data_addr := 16#28e + (#mode - 1) * 16#10;
               11..12: // Temperature
                   #mb_query.data_addr := 16#27e;
           END_CASE;
           #mb_query(data_ptr := #sign);
           #state += BOOL_TO_INT(#mb_query.Done);
       21: // Start use new coefficients.
           #mb_query(data_addr := 16#14c, data_ptr := #tDword);
           #state += BOOL_TO_INT(#mb_query.Done);
           // 22:
           //  #sign := #empty;
           // #state += 1;

           // =============

       30: // Chancel calibration
           #dword_14c := 0;
           #mb_query(data_addr := 16#14c, data_ptr := #dword_14c);
           #state += BOOL_TO_INT(#mb_query.Done);

           // =============

       ELSE // Reset
           #state := 0;
           #mode := 0;
           #Done := true;
           #error_cnt := 0;
   END_CASE;

   // Error handeling
   #error_cnt := BOOL_TO_USINT(#mb_query.Error);
   IF #ponsel_messure.sb.out.error
       OR #error_cnt > 3 // No more then x errors
   THEN
       #error_cnt := 0;
       #Error := true;
   END_IF;
END_FUNCTION_BLOCK

// ===== library: MasterCopy "ponselMesure_calibrateOksygen" =====

FUNCTION_BLOCK "ponselMesure_calibrateOksygen"   // FB2, SCL
{ S7_Optimized_Access := 'TRUE' }
VERSION : 0.1
   VAR_IN_OUT
      mb_query : "mb_query";
      ponsel_messure_oxygen : "Ponsel_mesure_Dissolved_oxygen";
   END_VAR
   VAR
      hmi : "ponselMesure_calibrateOxygenUdt";
      _ : Bool;
      state : Int;
      calibrate : "ponselMesure_calibrate";
   END_VAR
   VAR_TEMP
      empty : "ponselMesure_sign_udt";
   END_VAR
BEGIN
   CASE #state OF
       0:  // Wait for start signal.
           IF #hmi.startTempZeroCal THEN
               #calibrate.mode := 11; // Temperature zero (0 degrees C)
           ELSIF #hmi.startTempSpanCal THEN
               #calibrate.mode := 12; // Temperature span (25 degrees C)
           ELSIF #hmi.startOxygenZeroCal THEN
               #calibrate.mode := 1; // Oxygen zero (0 %)
           ELSIF #hmi.startOxygenSpanCal THEN
               #calibrate.mode := 4; // Oxygen span (100 %)
           ELSIF #hmi.save THEN
               #calibrate.state := 20; // Save changes.
           ELSIF #hmi.cancel THEN
               #calibrate.state := 30; // Cancel changes.
           END_IF;
           IF #calibrate.mode <> 0 THEN
               #calibrate.state := 10;
           END_IF;
           #state += 1;

       1:  // Wait for the calibration block.
           #calibrate(ref_value := #hmi.ref_value,
                      Done => #hmi.Done,
                      Error => #hmi.Error,
                      mb_query := #mb_query,
                      ponsel_messure := #ponsel_messure_oxygen.ponsel_mesure,
                      sign := #hmi.sign);
           IF #hmi.cancel THEN
               #calibrate.state := 30; // Cancel changes.
           ELSIF #calibrate.Done OR #mb_query.Error THEN
               #state := 0;
           END_IF;

   END_CASE;

   #hmi.cal_pending := #calibrate.dword_14c <> 0;

   #hmi.startTempZeroCal := false;
   #hmi.startTempSpanCal := false;
   #hmi.startOxygenZeroCal := false;
   #hmi.startOxygenSpanCal := false;
   #hmi.save := false;
   #hmi.cancel := false;
END_FUNCTION_BLOCK

// ===== library: MasterCopy "ponselMesure_calibrateOxygenUdt" =====

TYPE "ponselMesure_calibrateOxygenUdt"
   STRUCT
      startTempZeroCal : Bool;
      startTempSpanCal : Bool;
      startOxygenZeroCal : Bool;
      startOxygenSpanCal : Bool;
      save : Bool;
      cancel : Bool;
      ref_value : Real;
      sign : "ponselMesure_sign_udt";
      Done : Bool;
      Error : Bool;
      cal_pending : Bool;
   END_STRUCT;
END_TYPE

// ===== library: MasterCopy "ponselMesure_sign_udt" =====

TYPE "ponselMesure_sign_udt"
   STRUCT
      person : String[16];
      minute : String[2];
      hour : String[2];
      day : String[2];
      month : String[2];
      year : String[4];
      _ : String[4];
   END_STRUCT;
END_TYPE

(* ===== HMI "HMI_RT_2" =====
system functions are stored by id; their names below are inferred from use
connection "HMI_Connection_1": ETHERNET, S7_1200_OMS

HMI tags "Default tag table"
   "popupAnalogInTag" : WString[254] AT %DB1.DBX0.0

graphic list "@DiagnosticsStates": 0 '@Diagnostics_StateGood'; 1 '@Diagnostics_StateBad'

SlideinScreen "GraphX_Slidein_Left" 300x480
   Button "Button_4" at 43,212 size 190x34; TextOff 'Modbus'
      on Click: ActivateScreen("Modbus", 0)
   Button "Button_1" at 43,156 size 190x34; TextOff 'Home'
      on Click: ActivateScreen("Test", 0)
   Button "Button_2" at 43,268 size 190x34; TextOff 'Load balancer'
      on Click: ActivateScreen("load_balanser", 0)

SlideinScreen "GraphX_Slidein_Right" 267x480
   Button "Button_1" at 43,404 size 190x34; TextOff 'User mangement'
      on Click: ActivateScreen("UserMangement", 0)
   Button "Button_2" at 43,340 size 190x34; TextOff 'Diagnostics'
      on Click: ActivateScreen("Diagnostics", 0)
   Button "Button_3" at 43,276 size 190x34; TextOff 'Alarms'
      on Click: ActivateScreen("Alarms", 0)
   Button "Button_4" at 43,212 size 190x34; TextOff 'Test'
      on Click: ActivateScreen("Test", 0)